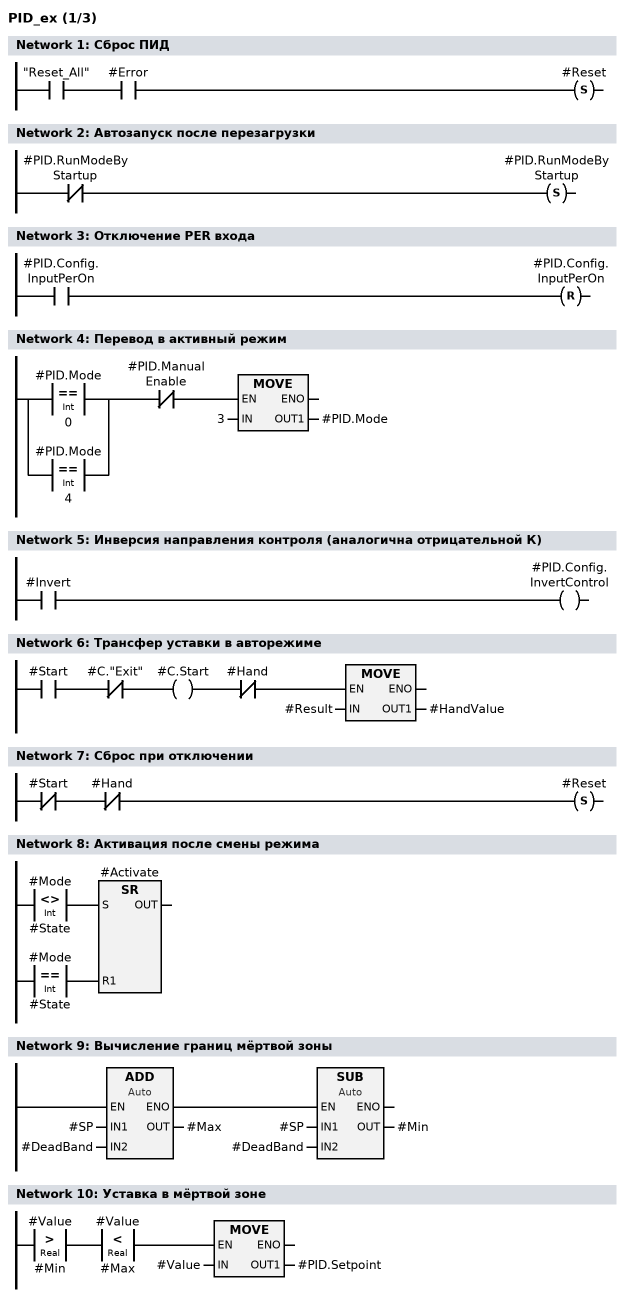
   RUNG wire#powerrail
      Contact( "Reset_All" )
      Contact( #Error )
      S_Coil( #Reset )
   END_RUNG
   // the same network as SCL:
   IF "Reset_All" AND #Error THEN #Reset := TRUE; END_IF;
END_REGION

REGION Network 2: Автозапуск после перезагрузки
   RUNG wire#powerrail
      I_Contact( #PID.RunModeByStartup )
      S_Coil( #PID.RunModeByStartup )
   END_RUNG
   // the same network as SCL:
   IF NOT #PID.RunModeByStartup THEN #PID.RunModeByStartup := TRUE; END_IF;
END_REGION

REGION Network 3: Отключение PER входа
   RUNG wire#powerrail
      Contact( #PID.Config.InputPerOn )
      R_Coil( #PID.Config.InputPerOn )
   END_RUNG
   // the same network as SCL:
   IF #PID.Config.InputPerOn THEN #PID.Config.InputPerOn := FALSE; END_IF;
END_REGION

REGION Network 4: Перевод в активный режим
   RUNG wire#powerrail
      { S7_Templates := "SrcType := Int" } EQ_Contact(in1 := #PID.Mode, in2 := 0)
      wire#w1
      I_Contact( #PID.ManualEnable )
      { S7_GenerateENO := "TRUE" } Move(in := 3, out1 => #PID.Mode)
   END_RUNG
   RUNG wire#powerrail
      { S7_Templates := "SrcType := Int" } EQ_Contact(in1 := #PID.Mode, in2 := 4)
   END_RUNG wire#w1
   // the same network as SCL:
   IF ((#PID.Mode = 0) OR (#PID.Mode = 4)) AND NOT #PID.ManualEnable THEN #PID.Mode := 3; END_IF;
END_REGION

REGION Network 5: Инверсия направления контроля (аналогична отрицательной К)
   RUNG wire#powerrail
      Contact( #Invert )
      Coil( #PID.Config.InvertControl )
   END_RUNG
   // the same network as SCL:
   #PID.Config.InvertControl := #Invert;
END_REGION

REGION Network 6: Трансфер уставки в авторежиме
   RUNG wire#powerrail
      Contact( #Start )
      I_Contact( #C."Exit" )
      Coil( #C.Start )
      I_Contact( #Hand )
      Move(in := #Result, out1 => #HandValue)
   END_RUNG
   // the same network as SCL:
   #C.Start := #Start AND NOT #C."Exit";
   IF #C.Start AND NOT #Hand THEN #HandValue := #Result; END_IF;
END_REGION

REGION Network 7: Сброс при отключении
   RUNG wire#powerrail
      I_Contact( #Start )
      I_Contact( #Hand )
      S_Coil( #Reset )
   END_RUNG
   // the same network as SCL:
   IF NOT #Start AND NOT #Hand THEN #Reset := TRUE; END_IF;
END_REGION

REGION Network 8: Активация после смены режима
   RUNG wire#powerrail
      { S7_Templates := "SrcType := Int" } NE_Contact(in1 := #Mode, in2 := #State)
      S_SR(operand := #Activate, r1 := wire#w1)
   END_RUNG
   RUNG wire#powerrail
      { S7_Templates := "SrcType := Int" } EQ_Contact(in1 := #Mode, in2 := #State)
   END_RUNG wire#w1
   // the same network as SCL:
   IF #Mode <> #State THEN
       #Activate := TRUE;   // SR flip-flop
   END_IF;
   IF #Mode = #State THEN #Activate := FALSE; END_IF;
END_REGION

REGION Network 9: Вычисление границ мёртвой зоны
   RUNG wire#powerrail
      Add(in1 := #SP, in2 := #DeadBand, out => #Max)
      Sub(in1 := #SP, in2 := #DeadBand, out => #Min)
   END_RUNG
   // the same network as SCL:
   #Max := #SP + #DeadBand;
   #Min := #SP - #DeadBand;
END_REGION

REGION Network 10: Уставка в мёртвой зоне
   RUNG wire#powerrail
      { S7_Templates := "SrcType := Real" } GT_Contact(in1 := #Value, in2 := #Min)
      { S7_Templates := "SrcType := Real" } LT_Contact(in1 := #Value, in2 := #Max)
      Move(in := #Value, out1 => #PID.Setpoint)
   END_RUNG
   // the same network as SCL:
   IF (#Value > #Min) AND (#Value < #Max) THEN #PID.Setpoint := #Value; END_IF;
END_REGION

REGION Network 11: Уставка вне мёртвой зоны
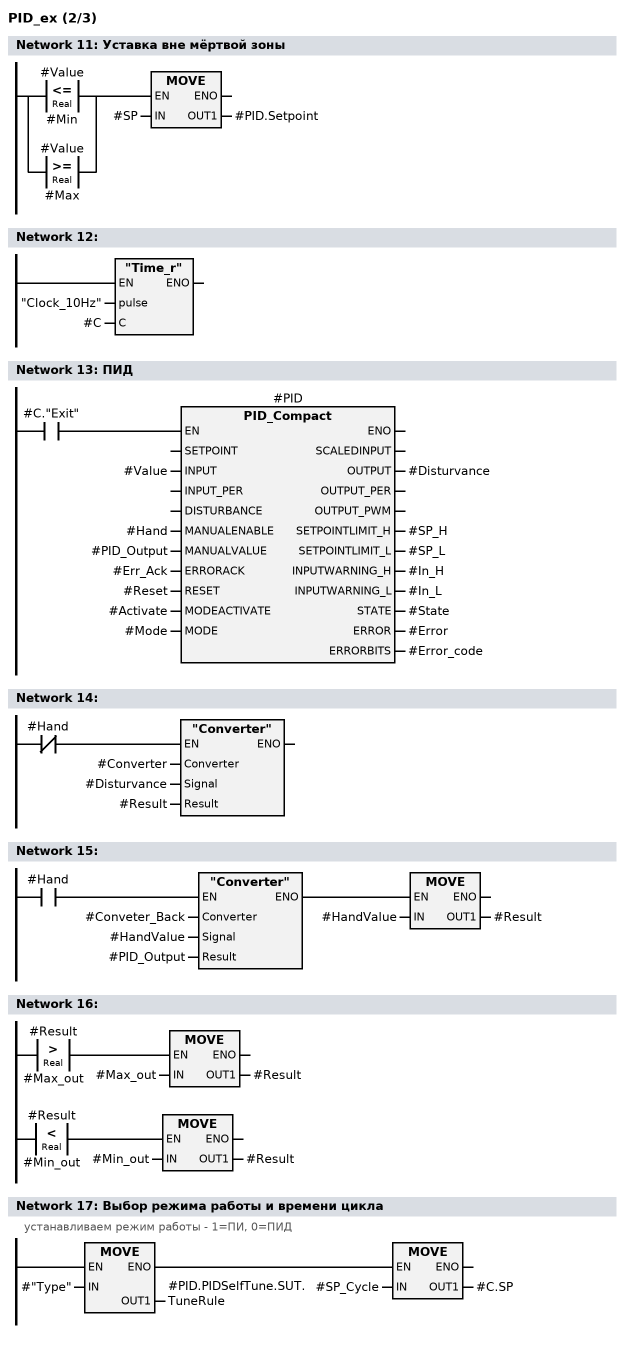
   RUNG wire#powerrail
      { S7_Templates := "SrcType := Real" } LE_Contact(in1 := #Value, in2 := #Min)
      wire#w1
      Move(in := #SP, out1 => #PID.Setpoint)
   END_RUNG
   RUNG wire#powerrail
      { S7_Templates := "SrcType := Real" } GE_Contact(in1 := #Value, in2 := #Max)
   END_RUNG wire#w1
   // the same network as SCL:
   IF (#Value <= #Min) OR (#Value >= #Max) THEN #PID.Setpoint := #SP; END_IF;
END_REGION

REGION Network 12
   RUNG wire#powerrail
      "Time_r"(pulse := "Clock_10Hz", C := #C)
   END_RUNG
   // the same network as SCL:
   "Time_r"(pulse := "Clock_10Hz", C := #C);
END_REGION

REGION Network 13: ПИД
   IF #C."Exit" THEN
       #PID(Input := #Value,   // PID_Compact
            ManualEnable := #Hand,
            ManualValue := #PID_Output,
            ErrorAck := #Err_Ack,
            Reset := #Reset,
            ModeActivate := #Activate,
            Mode := #Mode,
            Output => #Disturvance,
            SetpointLimit_H => #SP_H,
            SetpointLimit_L => #SP_L,
            InputWarning_H => #In_H,
            InputWarning_L => #In_L,
            State => #State,
            Error => #Error,
            ErrorBits => #Error_code);
   END_IF;
END_REGION

REGION Network 14
   RUNG wire#powerrail
      I_Contact( #Hand )
      "Converter"(Converter := #Converter, Signal := #Disturvance, Result := #Result)
   END_RUNG
   // the same network as SCL:
   IF NOT #Hand THEN "Converter"(Converter := #Converter, Signal := #Disturvance, Result := #Result); END_IF;
END_REGION

REGION Network 15
   RUNG wire#powerrail
      Contact( #Hand )
      "Converter"(Converter := #Conveter_Back, Signal := #HandValue, Result := #PID_Output)
      Move(in := #HandValue, out1 => #Result)
   END_RUNG
   // the same network as SCL:
   "Converter"(EN := #Hand,
               Converter := #Conveter_Back,
               Signal := #HandValue,
               Result := #PID_Output,
               ENO => #_w1);
   IF #_w1 THEN #Result := #HandValue; END_IF;
END_REGION

REGION Network 16
   RUNG wire#powerrail
      { S7_Templates := "SrcType := Real" } GT_Contact(in1 := #Result, in2 := #Max_out)
      Move(in := #Max_out, out1 => #Result)
   END_RUNG
   RUNG wire#powerrail
      { S7_Templates := "SrcType := Real" } LT_Contact(in1 := #Result, in2 := #Min_out)
      Move(in := #Min_out, out1 => #Result)
   END_RUNG
   // the same network as SCL:
   IF #Result > #Max_out THEN #Result := #Max_out; END_IF;
   IF #Result < #Min_out THEN #Result := #Min_out; END_IF;
END_REGION

REGION Network 17: Выбор режима работы и времени цикла
   // устанавливаем режим работы - 1=ПИ, 0=ПИД
   RUNG wire#powerrail
      { S7_GenerateENO := "TRUE" } Move(in := #"Type", out1 => #PID.PIDSelfTune.SUT.TuneRule)
      { S7_GenerateENO := "TRUE" } Move(in := #SP_Cycle, out1 => #C.SP)
   END_RUNG
   // the same network as SCL:
   // ENO of a box is taken as its EN; it also drops when the box reports an error
   #PID.PIDSelfTune.SUT.TuneRule := #"Type";
   #C.SP := #SP_Cycle;
END_REGION

REGION Network 18: Параметры регулирования
   // Задаём коэффициент пропорциональности и время интегрирования.
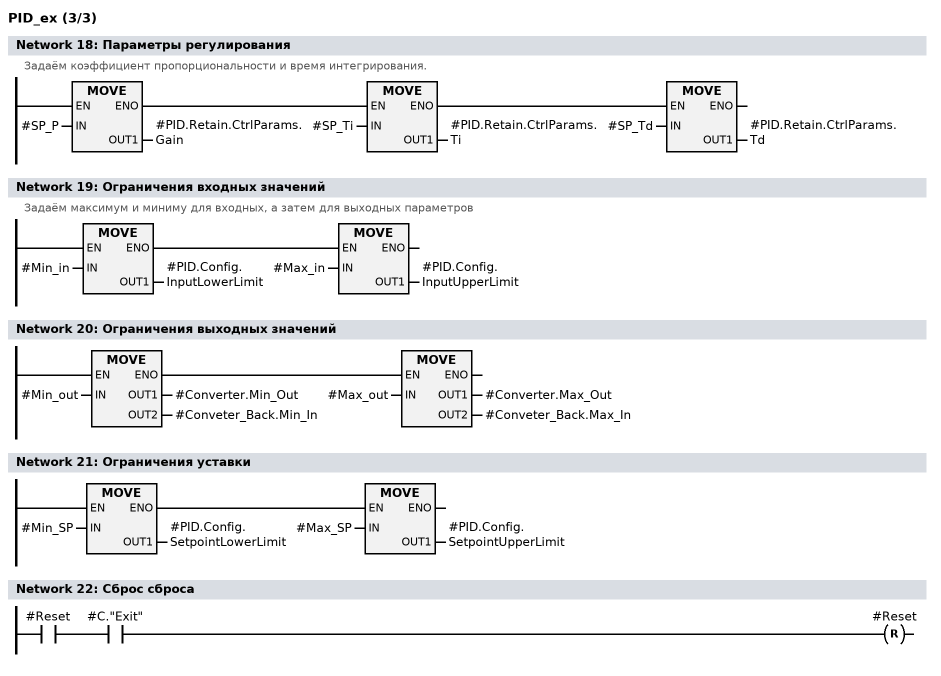
   RUNG wire#powerrail
      { S7_GenerateENO := "TRUE" } Move(in := #SP_P, out1 => #PID.Retain.CtrlParams.Gain)
      { S7_GenerateENO := "TRUE" } Move(in := #SP_Ti, out1 => #PID.Retain.CtrlParams.Ti)
      { S7_GenerateENO := "TRUE" } Move(in := #SP_Td, out1 => #PID.Retain.CtrlParams.Td)
   END_RUNG
   // the same network as SCL:
   // ENO of a box is taken as its EN; it also drops when the box reports an error
   #PID.Retain.CtrlParams.Gain := #SP_P;
   #PID.Retain.CtrlParams.Ti := #SP_Ti;
   #PID.Retain.CtrlParams.Td := #SP_Td;
END_REGION

REGION Network 19: Ограничения входных значений
   // Задаём максимум и миниму для входных, а затем для выходных параметров
   RUNG wire#powerrail
      { S7_GenerateENO := "TRUE" } Move(in := #Min_in, out1 => #PID.Config.InputLowerLimit)
      { S7_GenerateENO := "TRUE" } Move(in := #Max_in, out1 => #PID.Config.InputUpperLimit)
   END_RUNG
   // the same network as SCL:
   // ENO of a box is taken as its EN; it also drops when the box reports an error
   #PID.Config.InputLowerLimit := #Min_in;
   #PID.Config.InputUpperLimit := #Max_in;
END_REGION

REGION Network 20: Ограничения выходных значений
   RUNG wire#powerrail
      { S7_GenerateENO := "TRUE" } Move(in := #Min_out, out1 => #Converter.Min_Out, out2 => #Conveter_Back.Min_In)
      { S7_GenerateENO := "TRUE" } Move(in := #Max_out, out1 => #Converter.Max_Out, out2 => #Conveter_Back.Max_In)
   END_RUNG
   // the same network as SCL:
   // ENO of a box is taken as its EN; it also drops when the box reports an error
   #Converter.Min_Out := #Min_out;
   #Conveter_Back.Min_In := #Min_out;
   #Converter.Max_Out := #Max_out;
   #Conveter_Back.Max_In := #Max_out;
END_REGION

REGION Network 21: Ограничения уставки
   RUNG wire#powerrail
      { S7_GenerateENO := "TRUE" } Move(in := #Min_SP, out1 => #PID.Config.SetpointLowerLimit)
      { S7_GenerateENO := "TRUE" } Move(in := #Max_SP, out1 => #PID.Config.SetpointUpperLimit)
   END_RUNG
   // the same network as SCL:
   // ENO of a box is taken as its EN; it also drops when the box reports an error
   #PID.Config.SetpointLowerLimit := #Min_SP;
   #PID.Config.SetpointUpperLimit := #Max_SP;
END_REGION

REGION Network 22: Сброс сброса
   RUNG wire#powerrail
      Contact( #Reset )
      Contact( #C."Exit" )
      R_Coil( #Reset )
   END_RUNG
   // the same network as SCL:
   IF #Reset AND #C."Exit" THEN #Reset := FALSE; END_IF;
END_REGION
END_FUNCTION_BLOCK

FUNCTION "ASCII to Int" : Void   // FC12, LAD
{ S7_Optimized_Access := 'TRUE' }
VERSION : 0.1
   VAR_INPUT
      Code : Word;
   END_VAR
   VAR_OUTPUT
      Symbol : Int;
   END_VAR
BEGIN

REGION Network 1
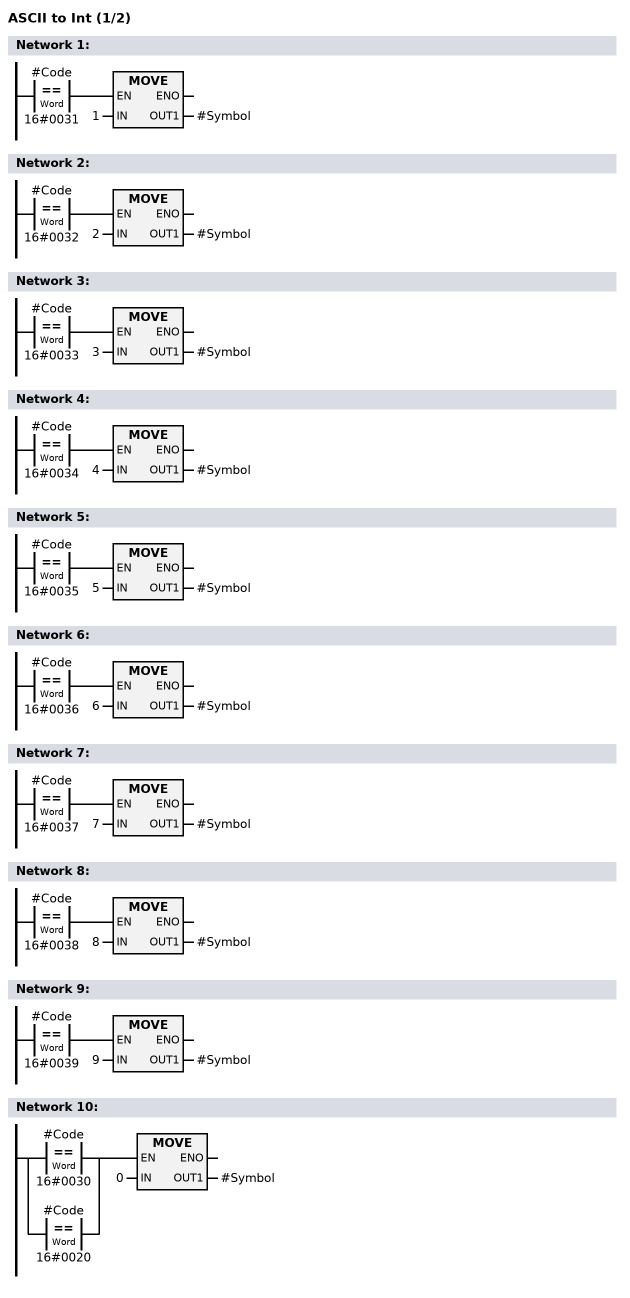
   RUNG wire#powerrail
      { S7_Templates := "SrcType := Word" } EQ_Contact(in1 := #Code, in2 := 16#0031)
      Move(in := 1, out1 => #Symbol)
   END_RUNG
   // the same network as SCL:
   IF #Code = 16#0031 THEN #Symbol := 1; END_IF;
END_REGION

REGION Network 2
   RUNG wire#powerrail
      { S7_Templates := "SrcType := Word" } EQ_Contact(in1 := #Code, in2 := 16#0032)
      Move(in := 2, out1 => #Symbol)
   END_RUNG
   // the same network as SCL:
   IF #Code = 16#0032 THEN #Symbol := 2; END_IF;
END_REGION

REGION Network 3
   RUNG wire#powerrail
      { S7_Templates := "SrcType := Word" } EQ_Contact(in1 := #Code, in2 := 16#0033)
      Move(in := 3, out1 => #Symbol)
   END_RUNG
   // the same network as SCL:
   IF #Code = 16#0033 THEN #Symbol := 3; END_IF;
END_REGION

REGION Network 4
   RUNG wire#powerrail
      { S7_Templates := "SrcType := Word" } EQ_Contact(in1 := #Code, in2 := 16#0034)
      Move(in := 4, out1 => #Symbol)
   END_RUNG
   // the same network as SCL:
   IF #Code = 16#0034 THEN #Symbol := 4; END_IF;
END_REGION

REGION Network 5
   RUNG wire#powerrail
      { S7_Templates := "SrcType := Word" } EQ_Contact(in1 := #Code, in2 := 16#0035)
      Move(in := 5, out1 => #Symbol)
   END_RUNG
   // the same network as SCL:
   IF #Code = 16#0035 THEN #Symbol := 5; END_IF;
END_REGION

REGION Network 6
   RUNG wire#powerrail
      { S7_Templates := "SrcType := Word" } EQ_Contact(in1 := #Code, in2 := 16#0036)
      Move(in := 6, out1 => #Symbol)
   END_RUNG
   // the same network as SCL:
   IF #Code = 16#0036 THEN #Symbol := 6; END_IF;
END_REGION

REGION Network 7
   RUNG wire#powerrail
      { S7_Templates := "SrcType := Word" } EQ_Contact(in1 := #Code, in2 := 16#0037)
      Move(in := 7, out1 => #Symbol)
   END_RUNG
   // the same network as SCL:
   IF #Code = 16#0037 THEN #Symbol := 7; END_IF;
END_REGION

REGION Network 8
   RUNG wire#powerrail
      { S7_Templates := "SrcType := Word" } EQ_Contact(in1 := #Code, in2 := 16#0038)
      Move(in := 8, out1 => #Symbol)
   END_RUNG
   // the same network as SCL:
   IF #Code = 16#0038 THEN #Symbol := 8; END_IF;
END_REGION

REGION Network 9
   RUNG wire#powerrail
      { S7_Templates := "SrcType := Word" } EQ_Contact(in1 := #Code, in2 := 16#0039)
      Move(in := 9, out1 => #Symbol)
   END_RUNG
   // the same network as SCL:
   IF #Code = 16#0039 THEN #Symbol := 9; END_IF;
END_REGION

REGION Network 10
   RUNG wire#powerrail
      { S7_Templates := "SrcType := Word" } EQ_Contact(in1 := #Code, in2 := 16#0030)
      wire#w1
      Move(in := 0, out1 => #Symbol)
   END_RUNG
   RUNG wire#powerrail
      { S7_Templates := "SrcType := Word" } EQ_Contact(in1 := #Code, in2 := 16#0020)
   END_RUNG wire#w1
   // the same network as SCL:
   IF (#Code = 16#0030) OR (#Code = 16#0020) THEN #Symbol := 0; END_IF;
END_REGION

REGION Network 11
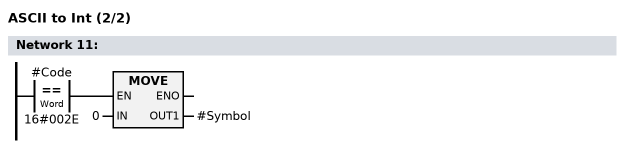
   RUNG wire#powerrail
      { S7_Templates := "SrcType := Word" } EQ_Contact(in1 := #Code, in2 := 16#002E)
      Move(in := 0, out1 => #Symbol)
   END_RUNG
   // the same network as SCL:
   IF #Code = 16#002E THEN #Symbol := 0; END_IF;
END_REGION
END_FUNCTION

FUNCTION "DRV_pulse" : Void   // FC100, LAD
{ S7_Optimized_Access := 'FALSE' }
VERSION : 0.1
   VAR_TEMP   // added for the SCL form of the ladder/FBD networks
      _w1 : Bool;
      _w2 : Bool;
   END_VAR
BEGIN

REGION Network 1
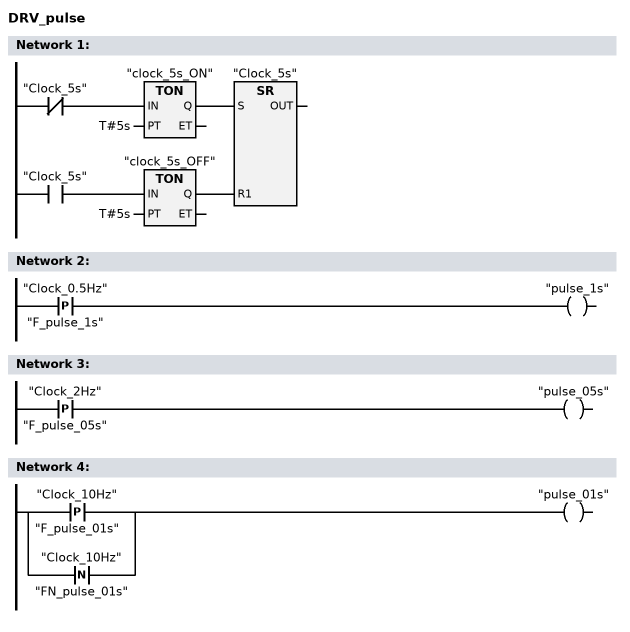
   "clock_5s_ON".TON(IN := NOT "Clock_5s", PT := T#5s);
   "clock_5s_OFF".TON(IN := "Clock_5s", PT := T#5s);
   IF "clock_5s_ON".Q THEN
       "Clock_5s" := TRUE;   // SR flip-flop
   END_IF;
   IF "clock_5s_OFF".Q THEN "Clock_5s" := FALSE; END_IF;
END_REGION

REGION Network 2
   RUNG wire#powerrail
      P_Contact(operand := "Clock_0.5Hz", bit := "F_pulse_1s")
      Coil( "pulse_1s" )
   END_RUNG
   // the same network as SCL:
   #_w1 := "Clock_0.5Hz" AND NOT "F_pulse_1s";   // rising edge of "Clock_0.5Hz"
   "F_pulse_1s" := "Clock_0.5Hz";
   "pulse_1s" := #_w1;
END_REGION

REGION Network 3
   RUNG wire#powerrail
      P_Contact(operand := "Clock_2Hz", bit := "F_pulse_05s")
      Coil( "pulse_05s" )
   END_RUNG
   // the same network as SCL:
   #_w1 := "Clock_2Hz" AND NOT "F_pulse_05s";   // rising edge of "Clock_2Hz"
   "F_pulse_05s" := "Clock_2Hz";
   "pulse_05s" := #_w1;
END_REGION

REGION Network 4
   RUNG wire#powerrail
      P_Contact(operand := "Clock_10Hz", bit := "F_pulse_01s")
      wire#w1
      Coil( "pulse_01s" )
   END_RUNG
   RUNG wire#powerrail
      N_Contact(operand := "Clock_10Hz", bit := "FN_pulse_01s")
   END_RUNG wire#w1
   // the same network as SCL:
   #_w1 := "Clock_10Hz" AND NOT "F_pulse_01s";   // rising edge of "Clock_10Hz"
   "F_pulse_01s" := "Clock_10Hz";
   #_w2 := NOT "Clock_10Hz" AND "FN_pulse_01s";   // falling edge of "Clock_10Hz"
   "FN_pulse_01s" := "Clock_10Hz";
   "pulse_01s" := #_w1 OR #_w2;
END_REGION
END_FUNCTION

FUNCTION "DRV_End" : Void   // FC101, LAD
{ S7_Optimized_Access := 'TRUE' }
VERSION : 0.1
BEGIN

REGION Network 1: Одно из устройств нижнего уровня в ручном режиме
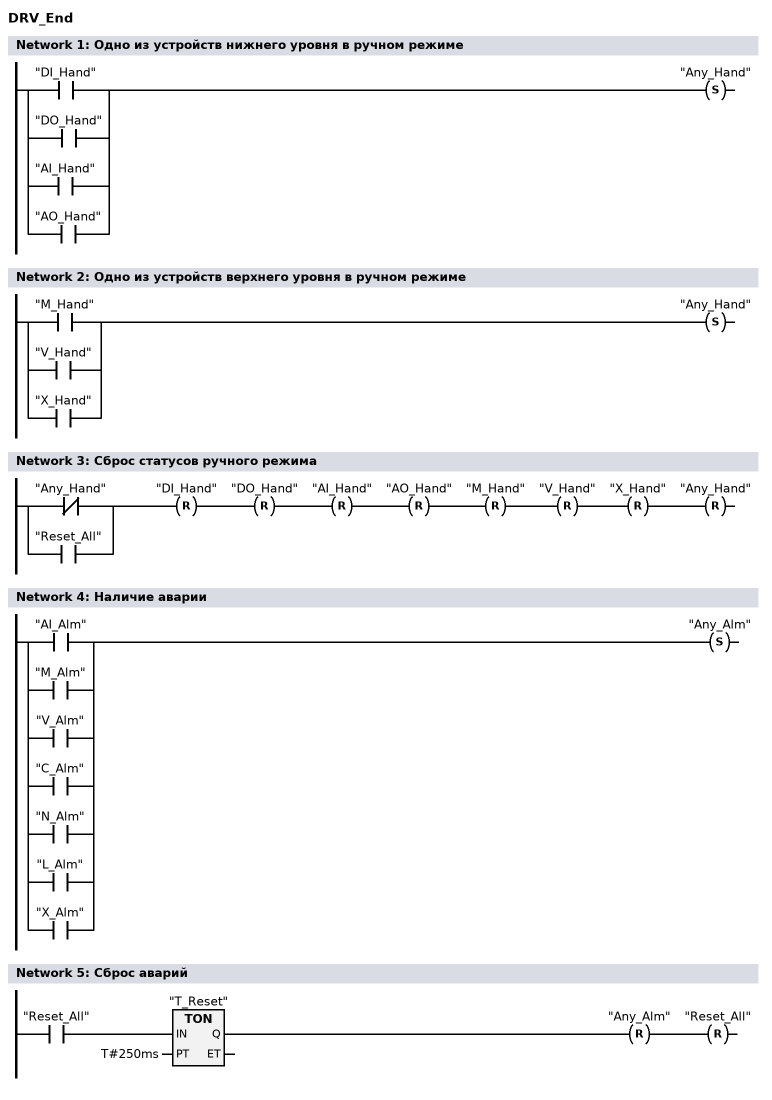
   RUNG wire#powerrail
      Contact( "DI_Hand" )
      wire#w1
      S_Coil( "Any_Hand" )
   END_RUNG
   RUNG wire#powerrail
      Contact( "DO_Hand" )
   END_RUNG wire#w1
   RUNG wire#powerrail
      Contact( "AI_Hand" )
   END_RUNG wire#w1
   RUNG wire#powerrail
      Contact( "AO_Hand" )
   END_RUNG wire#w1
   // the same network as SCL:
   IF "DI_Hand" OR "DO_Hand" OR "AI_Hand" OR "AO_Hand" THEN "Any_Hand" := TRUE; END_IF;
END_REGION

REGION Network 2: Одно из устройств верхнего уровня в ручном режиме
   RUNG wire#powerrail
      Contact( "M_Hand" )
      wire#w1
      S_Coil( "Any_Hand" )
   END_RUNG
   RUNG wire#powerrail
      Contact( "V_Hand" )
   END_RUNG wire#w1
   RUNG wire#powerrail
      Contact( "X_Hand" )
   END_RUNG wire#w1
   // the same network as SCL:
   IF "M_Hand" OR "V_Hand" OR "X_Hand" THEN "Any_Hand" := TRUE; END_IF;
END_REGION

REGION Network 3: Сброс статусов ручного режима
   RUNG wire#powerrail
      I_Contact( "Any_Hand" )
      wire#w1
      R_Coil( "DI_Hand" )
      R_Coil( "DO_Hand" )
      R_Coil( "AI_Hand" )
      R_Coil( "AO_Hand" )
      R_Coil( "M_Hand" )
      R_Coil( "V_Hand" )
      R_Coil( "X_Hand" )
      R_Coil( "Any_Hand" )
   END_RUNG
   RUNG wire#powerrail
      Contact( "Reset_All" )
   END_RUNG wire#w1
   // the same network as SCL:
   IF NOT "Any_Hand" OR "Reset_All" THEN
       "DI_Hand" := FALSE;
       "DO_Hand" := FALSE;
       "AI_Hand" := FALSE;
       "AO_Hand" := FALSE;
       "M_Hand" := FALSE;
       "V_Hand" := FALSE;
       "X_Hand" := FALSE;
       "Any_Hand" := FALSE;
   END_IF;
END_REGION

REGION Network 4: Наличие аварии
   RUNG wire#powerrail
      Contact( "AI_Alm" )
      wire#w1
      S_Coil( "Any_Alm" )
   END_RUNG
   RUNG wire#powerrail
      Contact( "M_Alm" )
   END_RUNG wire#w1
   RUNG wire#powerrail
      Contact( "V_Alm" )
   END_RUNG wire#w1
   RUNG wire#powerrail
      Contact( "C_Alm" )
   END_RUNG wire#w1
   RUNG wire#powerrail
      Contact( "N_Alm" )
   END_RUNG wire#w1
   RUNG wire#powerrail
      Contact( "L_Alm" )
   END_RUNG wire#w1
   RUNG wire#powerrail
      Contact( "X_Alm" )
   END_RUNG wire#w1
   // the same network as SCL:
   IF "AI_Alm" OR "M_Alm" OR "V_Alm" OR "C_Alm" OR "N_Alm" OR "L_Alm" OR "X_Alm" THEN
       "Any_Alm" := TRUE;
   END_IF;
END_REGION

REGION Network 5: Сброс аварий
   "T_Reset".TON(IN := "Reset_All", PT := T#250ms);
   IF "T_Reset".Q THEN
       "Any_Alm" := FALSE;
       "Reset_All" := FALSE;
   END_IF;
END_REGION
END_FUNCTION

FUNCTION "Converter" : Void   // FC102, LAD
TITLE = Драйвер линеаризации аналогового сигнала
{ S7_Optimized_Access := 'FALSE' }
VERSION : 0.1
   VAR_INPUT
      Converter : Struct
         Use_Min_In : Bool;   // Отсекать входные значения ниже минимума
         Use_Max_In : Bool;   // Отсекать входные значения выше максимума
         Use_Min_Out : Bool;   // Отсекать результат ниже минимума
         Use_Max_Out : Bool;   // Отсекать результат выше максимума
         IO : Bool;   // Входной/Выходной режим
         Inverse : Bool;   // Инверсия выхода
         Min_In : Real;   // Минимальный входной сигнал
         Max_In : Real;   // Максимальный входной сигнал
         Min_Out : Real;   // Минимальный выходной сигнал
         Max_Out : Real;   // Максимальный выходной сигнал
      END_STRUCT;
   END_VAR
   VAR_IN_OUT
      Signal : Real;   // Входной сигнал
      Result : Real;   // Результат линеаризации
   END_VAR
   VAR_TEMP
      Range_In : Real;   // Диапазон входного сигнала
      Range_Out : Real;   // Диапазон выходного сигнала
      T_T : Real;   // Соотношение диапазонов
      R_Sig : Real;   // Поправка на отрицательные значения
   END_VAR
BEGIN

REGION Network 1: Проверка нижнего уровня входного сигнала
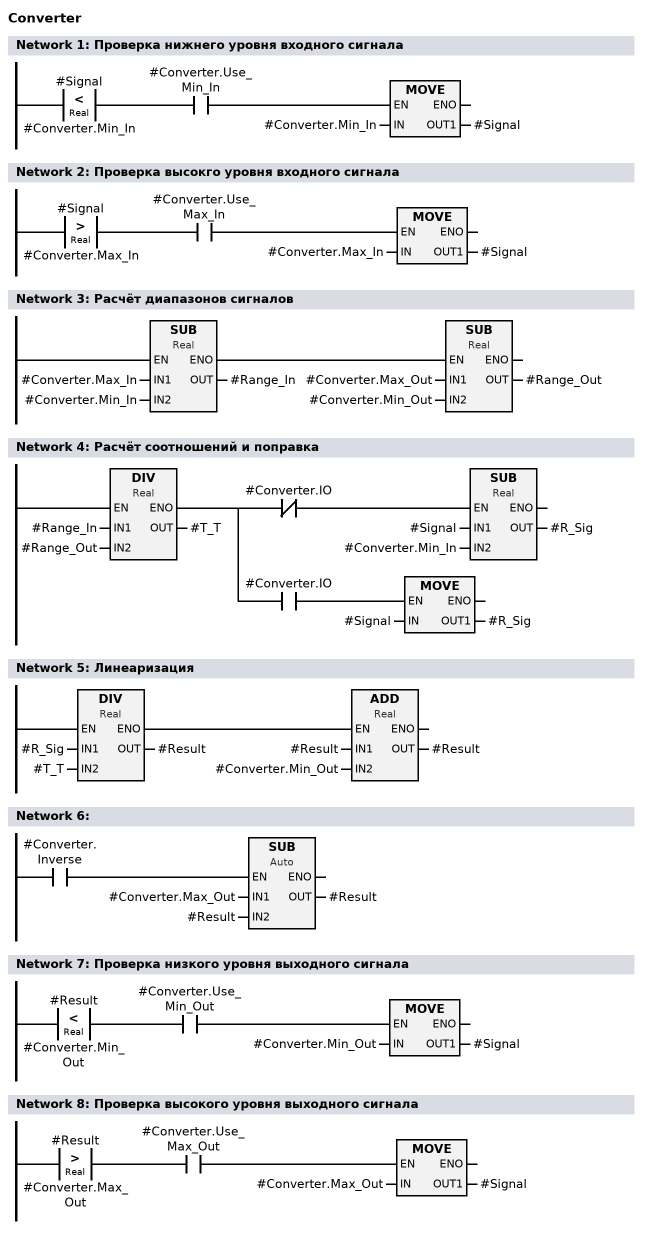
   RUNG wire#powerrail
      { S7_Templates := "SrcType := Real" } LT_Contact(in1 := #Signal, in2 := #Converter.Min_In)
      Contact( #Converter.Use_Min_In )
      Move(in := #Converter.Min_In, out1 => #Signal)
   END_RUNG
   // the same network as SCL:
   IF (#Signal < #Converter.Min_In) AND #Converter.Use_Min_In THEN #Signal := #Converter.Min_In; END_IF;
END_REGION

REGION Network 2: Проверка высокго уровня входного сигнала
   RUNG wire#powerrail
      { S7_Templates := "SrcType := Real" } GT_Contact(in1 := #Signal, in2 := #Converter.Max_In)
      Contact( #Converter.Use_Max_In )
      Move(in := #Converter.Max_In, out1 => #Signal)
   END_RUNG
   // the same network as SCL:
   IF (#Signal > #Converter.Max_In) AND #Converter.Use_Max_In THEN #Signal := #Converter.Max_In; END_IF;
END_REGION

REGION Network 3: Расчёт диапазонов сигналов
   RUNG wire#powerrail
      { S7_Templates := "SrcType := Real"; S7_GenerateENO := "TRUE" } Sub(in1 := #Converter.Max_In, in2 := #Converter.Min_In, out => #Range_In)
      { S7_Templates := "SrcType := Real"; S7_GenerateENO := "TRUE" } Sub(in1 := #Converter.Max_Out, in2 := #Converter.Min_Out, out => #Range_Out)
   END_RUNG
   // the same network as SCL:
   // ENO of a box is taken as its EN; it also drops when the box reports an error
   #Range_In := #Converter.Max_In - #Converter.Min_In;
   #Range_Out := #Converter.Max_Out - #Converter.Min_Out;
END_REGION

REGION Network 4: Расчёт соотношений и поправка
   RUNG wire#powerrail
      { S7_Templates := "SrcType := Real"; S7_GenerateENO := "TRUE" } Div(in1 := #Range_In, in2 := #Range_Out, out => #T_T)
      wire#w1
      I_Contact( #Converter.IO )
      { S7_Templates := "SrcType := Real"; S7_GenerateENO := "TRUE" } Sub(in1 := #Signal, in2 := #Converter.Min_In, out => #R_Sig)
   END_RUNG
   RUNG wire#w1
      Contact( #Converter.IO )
      Move(in := #Signal, out1 => #R_Sig)
   END_RUNG
   // the same network as SCL:
   // ENO of a box is taken as its EN; it also drops when the box reports an error
   #T_T := #Range_In / #Range_Out;
   IF NOT #Converter.IO THEN #R_Sig := #Signal - #Converter.Min_In; END_IF;
   IF #Converter.IO THEN #R_Sig := #Signal; END_IF;
END_REGION

REGION Network 5: Линеаризация
   RUNG wire#powerrail
      { S7_Templates := "SrcType := Real"; S7_GenerateENO := "TRUE" } Div(in1 := #R_Sig, in2 := #T_T, out => #Result)
      { S7_Templates := "SrcType := Real"; S7_GenerateENO := "TRUE" } Add(in1 := #Result, in2 := #Converter.Min_Out, out => #Result)
   END_RUNG
   // the same network as SCL:
   // ENO of a box is taken as its EN; it also drops when the box reports an error
   #Result := #R_Sig / #T_T;
   #Result := #Result + #Converter.Min_Out;
END_REGION

REGION Network 6
   RUNG wire#powerrail
      Contact( #Converter.Inverse )
      Sub(in1 := #Converter.Max_Out, in2 := #Result, out => #Result)
   END_RUNG
   // the same network as SCL:
   IF #Converter.Inverse THEN #Result := #Converter.Max_Out - #Result; END_IF;
END_REGION

REGION Network 7: Проверка низкого уровня выходного сигнала
   RUNG wire#powerrail
      { S7_Templates := "SrcType := Real" } LT_Contact(in1 := #Result, in2 := #Converter.Min_Out)
      Contact( #Converter.Use_Min_Out )
      Move(in := #Converter.Min_Out, out1 => #Signal)
   END_RUNG
   // the same network as SCL:
   IF (#Result < #Converter.Min_Out) AND #Converter.Use_Min_Out THEN #Signal := #Converter.Min_Out; END_IF;
END_REGION

REGION Network 8: Проверка высокого уровня выходного сигнала
   RUNG wire#powerrail
      { S7_Templates := "SrcType := Real" } GT_Contact(in1 := #Result, in2 := #Converter.Max_Out)
      Contact( #Converter.Use_Max_Out )
      Move(in := #Converter.Max_Out, out1 => #Signal)
   END_RUNG
   // the same network as SCL:
   IF (#Result > #Converter.Max_Out) AND #Converter.Use_Max_Out THEN #Signal := #Converter.Max_Out; END_IF;
END_REGION
END_FUNCTION

FUNCTION "Balancer" : Void   // FC103, LAD
TITLE = Балансировка нагрузки двух устройств по наработке и аварии
{ S7_Optimized_Access := 'FALSE' }